   GraphicIOField "PlotLight_Round_G_33" at 416,264 size 24x24; PictureOn "PilotLight_Round_G_On_256c"; PictureOff "PilotLight_Round_G_Off_256c"
      ProcessValue <- "Senzor 2 proximitate softstarter aer destacker"

screen "Manual.Stacker" 800x480, template "TemplateWithClockAndBackBtnForManual"
   on GenerateScreen: SetBit("Maintenance")
   on ClearScreen: ResetBit("Maintenance")
   TextField "Text field_14" at 494,54 size 179x20; Text 'Comanda 1 softstarter aer'
   TextField "Text field_15" at 494,134 size 190x20; Text 'Comanda cilindru vertical jos'
   TextField "Text field_16" at 494,174 size 193x20; Text 'Comanda cilindru vertical sus'
   TextField "Text field_17" at 494,214 size 155x20; Text 'Comanda furca retrasa'
   TextField "Text field_18" at 494,254 size 153x20; Text 'Comanda furca extinsa'
   Switch "Switch_1" at 696,128 size 64x32; CaptionText 'Switch'; TextOff 'OFF'; TextOn 'ON'
      ProcessValue <- "S_Comanda cilindru vertical jos"
      on SwitchOn: SetBit("S_Comanda cilindru vertical jos")
      on SwitchOff: ResetBit("S_Comanda cilindru vertical jos")
   GraphicIOField "PlotLight_Round_G_2" at 160,48 size 24x24; PictureOff "PilotLight_Round_G_Off_256c"; PictureOn "PilotLight_Round_G_On_256c"
      ProcessValue <- "DB_PalletDispenser_PD2_Stacking_DB_PD1_MiddlePosition"
   TextField "Text field_3" at 16,50 size 126x20; Text 'PD1 MiddlePosition'
   Switch "Switch_2" at 696,48 size 64x32; CaptionText 'Switch'; TextOff 'OFF'; TextOn 'ON'
      ProcessValue <- "Comanda 1 softstarter aer stacker"
      on SwitchOn: SetBit("Comanda 1 softstarter aer stacker")
      on SwitchOff: ResetBit("Comanda 1 softstarter aer stacker")
   Switch "Switch_3" at 696,168 size 64x32; CaptionText 'Switch'; TextOff 'OFF'; TextOn 'ON'
      ProcessValue <- "S_Comanda cilindru vertical sus"
      on SwitchOn: SetBit("S_Comanda cilindru vertical sus")
      on SwitchOff: ResetBit("S_Comanda cilindru vertical sus")
   Switch "Switch_4" at 696,208 size 64x32; CaptionText 'Switch'; TextOff 'OFF'; TextOn 'ON'
      ProcessValue <- "S_Comanda furca retrasa"
      on SwitchOn: SetBit("S_Comanda furca retrasa")
      on SwitchOff: ResetBit("S_Comanda furca retrasa")
   Switch "Switch_5" at 696,248 size 64x32; CaptionText 'Switch'; TextOff 'OFF'; TextOn 'ON'
      ProcessValue <- "S_Comanda furca extinsa"
      on SwitchOn: SetBit("S_Comanda furca extinsa")
      on SwitchOff: ResetBit("S_Comanda furca extinsa")
   TextField "Text field_21" at 494,94 size 179x20; Text 'Comanda 2 softstarter aer'
   Switch "Switch_8" at 696,88 size 64x32; CaptionText 'Switch'; TextOff 'OFF'; TextOn 'ON'
      ProcessValue <- "Comanda 2 softstarter aer stacker"
      on SwitchOn: SetBit("Comanda 2 softstarter aer stacker")
      on SwitchOff: ResetBit("Comanda 2 softstarter aer stacker")
   GraphicIOField "PlotLight_Round_G_1" at 160,72 size 24x24; PictureOn "PilotLight_Round_G_On_256c"; PictureOff "PilotLight_Round_G_Off_256c"
      ProcessValue <- "DB_PalletDispenser_PD2_Stacking_DB_PD1_Up"
   TextField "Text field_1" at 16,74 size 50x20; Text 'PD1 Up'
   GraphicIOField "PlotLight_Round_G_3" at 160,96 size 24x24; PictureOn "PilotLight_Round_G_On_256c"; PictureOff "PilotLight_Round_G_Off_256c"
      ProcessValue <- "DB_PalletDispenser_PD2_Stacking_DB_PD1_Down"
   TextField "Text field_2" at 16,98 size 70x20; Text 'PD1 Down'
   GraphicIOField "PlotLight_Round_G_4" at 160,120 size 24x24; PictureOn "PilotLight_Round_G_On_256c"; PictureOff "PilotLight_Round_G_Off_256c"
      ProcessValue <- "DB_PalletDispenser_PD2_Stacking_DB_PD1_Forks_In"
   TextField "Text field_4" at 16,122 size 85x20; Text 'PD1 Forks In'
   GraphicIOField "PlotLight_Round_G_5" at 160,144 size 24x24; PictureOff "PilotLight_Round_G_Off_256c"; PictureOn "PilotLight_Round_G_On_256c"
      ProcessValue <- "DB_PalletDispenser_PD2_Stacking_DB_PD1_Forks_Out"
   TextField "Text field_5" at 16,146 size 95x20; Text 'PD1 Forks Out'
   GraphicIOField "PlotLight_Round_G_7" at 160,168 size 24x24; PictureOn "PilotLight_Round_G_On_256c"; PictureOff "PilotLight_Round_G_Off_256c"
      ProcessValue <- "DB_PalletDispenser_PD2_Stacking_DB_Alarm_Active"
   TextField "Text field_7" at 16,170 size 89x20; Text 'Alarm Active'
   GraphicIOField "PlotLight_Round_G_8" at 416,48 size 24x24; PictureOff "PilotLight_Round_G_Off_256c"; PictureOn "PilotLight_Round_G_On_256c"
      ProcessValue <- "S_Cilindru extins"
   TextField "Text field_8" at 240,50 size 111x20; Text 'S_Cilindru extins'
   GraphicIOField "PlotLight_Round_G_9" at 416,72 size 24x24; PictureOff "PilotLight_Round_G_Off_256c"; PictureOn "PilotLight_Round_G_On_256c"
      ProcessValue <- "S_Cilindru retras"
   TextField "Text field_9" at 240,74 size 113x20; Text 'S_Cilindru retras'
   GraphicIOField "PlotLight_Round_G_10" at 416,96 size 24x24; PictureOn "PilotLight_Round_G_On_256c"; PictureOff "PilotLight_Round_G_Off_256c"
      ProcessValue <- "S_Cilindru vertical jos"
   TextField "Text field_10" at 240,98 size 144x20; Text 'S_Cilindru vertical jos'
   GraphicIOField "PlotLight_Round_G_11" at 416,120 size 24x24; PictureOn "PilotLight_Round_G_On_256c"; PictureOff "PilotLight_Round_G_Off_256c"
      ProcessValue <- "S_Cilindru vertical mijloc"
   TextField "Text field_11" at 240,122 size 161x20; Text 'S_Cilindru vertical mijloc'
   GraphicIOField "PlotLight_Round_G_12" at 416,144 size 24x24; PictureOn "PilotLight_Round_G_On_256c"; PictureOff "PilotLight_Round_G_Off_256c"
      ProcessValue <- "S_Cilindru vertical sus"
   TextField "Text field_12" at 240,146 size 147x20; Text 'S_Cilindru vertical sus'
   GraphicIOField "PlotLight_Round_G_13" at 416,168 size 24x24; PictureOff "PilotLight_Round_G_Off_256c"; PictureOn "PilotLight_Round_G_On_256c"
      ProcessValue <- "S_Lungime 1"
   TextField "Text field_13" at 240,170 size 86x20; Text 'S_Lungime 1'
   GraphicIOField "PlotLight_Round_G_14" at 416,192 size 24x24; PictureOff "PilotLight_Round_G_Off_256c"; PictureOn "PilotLight_Round_G_On_256c"
      ProcessValue <- "S_Lungime 2"
   TextField "Text field_19" at 240,194 size 86x20; Text 'S_Lungime 2'
   GraphicIOField "PlotLight_Round_G_15" at 416,216 size 24x24; PictureOn "PilotLight_Round_G_On_256c"; PictureOff "PilotLight_Round_G_Off_256c"
      ProcessValue <- "S_Lungime 3"
   TextField "Text field_20" at 240,218 size 86x20; Text 'S_Lungime 3'
   GraphicIOField "PlotLight_Round_G_6" at 416,240 size 24x24; PictureOff "PilotLight_Round_G_Off_256c"; PictureOn "PilotLight_Round_G_On_256c"
      ProcessValue <- "S_Detectie palet"
   TextField "Text field_6" at 240,242 size 113x20; Text 'S_Detectie palet'
   GraphicIOField "PlotLight_Round_G_30" at 416,264 size 24x24; PictureOn "PilotLight_Round_G_On_256c"; PictureOff "PilotLight_Round_G_Off_256c"
      ProcessValue <- "Senzor 1 proximitate softstarter aer stacker"
   TextField "Text field_31" at 112,266 size 296x20; Text 'Senzor 1 proximitate softstarter aer stacker'
   GraphicIOField "PlotLight_Round_G_34" at 416,288 size 24x24; PictureOn "PilotLight_Round_G_On_256c"; PictureOff "PilotLight_Round_G_Off_256c"
      ProcessValue <- "Senzor 2 proximitate softstarter aer stacker"
   TextField "Text field_35" at 112,290 size 296x20; Text 'Senzor 2 proximitate softstarter aer stacker'

Template "TemplateWithClock" 800x480
   DateTimeField "Template_Date/time field_1" at 624,10 size 172x21
   GraphicView "Template_Graphic view_1" at 592,384 size 208x96; Picture "energom logo gonzales_1"

Template "TemplateWithClockAndBackBtn" 800x480
   Button "SB_NavigateLeft_48x48" at 72,0 size 64x40; TextOff 'Text'; PictureOff "SB_NavigateLeft_48x48_256c"
      on Press: function_efd93a16()
   Button "SB_NavigateHome_48x48" at 0,0 size 64x40; TextOff 'Text'; PictureOff "SB_NavigateHome_48x48_256c"
      on Press: ActivateScreen("Main", 0)
   DateTimeField "Template_Date/time field_1" at 624,10 size 172x21
   GraphicView "Template_Graphic view_1" at 592,384 size 208x96; Picture "energom logo gonzales_1"

Template "TemplateWithClockAndBackBtnForStatistics" 800x480
   Button "SB_NavigateHome_48x48" at 0,0 size 64x40; TextOff 'Text'; PictureOff "SB_NavigateHome_48x48_256c"
      on Press: ActivateScreen("Main", 0)
   Button "Button_4" at 8,392 size 136x80; TextOff 'Paleti Reparati'; Authorization "Operate"
      on Press: ActivateScreen("Production.Repair", 0); SetTag("CurrentScreenStatistics", 0)
      Visibility <- "CurrentUserGroup"
      Appearance <- "CurrentScreenStatistics"
   Button "Button_1" at 152,392 size 136x80; TextOff 'Paleti Demontati'; Authorization "Operate"
      on Press: ActivateScreen("Production.Destroy", 0); SetTag("CurrentScreenStatistics", 1)
      Visibility <- "CurrentUserGroup"
      Appearance <- "CurrentScreenStatistics"
   Button "Button_2" at 296,392 size 136x80; TextOff 'Energie'; Authorization "Operate"
      on Press: ActivateScreen("Energy", 0); SetTag("CurrentScreenStatistics", 2)
      Visibility <- "CurrentUserGroup"
      Appearance <- "CurrentScreenStatistics"
   Button "Button_3" at 440,392 size 136x80; TextOff 'Protectii'; Authorization "Operate"
      on Press: ActivateScreen("Safety", 0); SetTag("CurrentScreenStatistics", 3)
      Visibility <- "CurrentUserGroup"
      Appearance <- "CurrentScreenStatistics"
   DateTimeField "Template_Date/time field_1" at 624,10 size 172x21
   GraphicView "Template_Graphic view_1" at 592,384 size 208x96; Picture "energom logo gonzales_1"

Template "TemplateWithClockAndBackBtnForManual" 800x480
   Button "SB_NavigateHome_48x48" at 0,0 size 64x40; TextOff 'Text'; PictureOff "SB_NavigateHome_48x48_256c"
      on Press: ActivateScreen("Main", 0)
   DateTimeField "Template_Date/time field_1" at 624,10 size 172x21
   Button "Button_5" at 8,392 size 136x36; TextOff 'General'; Authorization "Operate"
      on Press: ActivateScreen("Manual.General", 0); SetTag("CurrentScreenManual", 0)
      Visibility <- "CurrentUserGroup"
      Appearance <- "CurrentScreenManual"
   Button "Button_6" at 152,392 size 136x36; TextOff 'Destacker'; Authorization "Operate"
      on Press: ActivateScreen("Manual.Destacker", 0); SetTag("CurrentScreenManual", 2)
      Visibility <- "CurrentUserGroup"
      Appearance <- "CurrentScreenManual"
   Button "Button_7" at 296,392 size 136x36; TextOff 'Stacker'; Authorization "Operate"
      on Press: ActivateScreen("Manual.Stacker", 0); SetTag("CurrentScreenManual", 4)
      Visibility <- "CurrentUserGroup"
      Appearance <- "CurrentScreenManual"
   Button "Button_8" at 8,436 size 136x36; TextOff 'Safety'; Authorization "Operate"
      on Press: ActivateScreen("Manual.Safety", 0); SetTag("CurrentScreenManual", 1)
      Visibility <- "CurrentUserGroup"
      Appearance <- "CurrentScreenManual"
   Button "Button_1" at 440,392 size 136x36; TextOff 'Transfer'; Authorization "Operate"
      on Press: ActivateScreen("Manual.Transfer", 0); SetTag("CurrentScreenManual", 6)
      Visibility <- "CurrentUserGroup"
      Appearance <- "CurrentScreenManual"
   GraphicView "Template_Graphic view_1" at 592,384 size 208x96; Picture "energom logo gonzales_1"
   Button "Button_2" at 152,436 size 136x36; TextOff 'Conveioare Destacker'; Authorization "Operate"
      on Press: ActivateScreen("Manual.DestackerConveyors", 0); SetTag("CurrentScreenManual", 3)
      Visibility <- "CurrentUserGroup"
      Appearance <- "CurrentScreenManual"
   Button "Button_3" at 296,436 size 136x36; TextOff 'Conveioare Stacker'; Authorization "Operate"
      on Press: ActivateScreen("Manual.StackerConveyors", 0); SetTag("CurrentScreenManual", 5)
      Visibility <- "CurrentUserGroup"
      Appearance <- "CurrentScreenManual"
   Button "Button_4" at 440,436 size 136x36; TextOff 'Diagnoza IO Link'; Authorization "Operate"
      on Press: ActivateScreen("Manual.IOLinkDiag", 0); SetTag("CurrentScreenManual", 7)
      Visibility <- "CurrentUserGroup"
      Appearance <- "CurrentScreenManual"

scheduled task "ChangeUserTask"
   on Action: function_f41c6f6c("CurrentUser"); function_e1ab61de("CurrentUserGroup"); function_de9337da()
*)

(* ===== HMI "HMI_RT_1" =====

graphic list "List": 1 'Graphic_4'; 2 'Graphic_6'; 4..16 'Graphic_7'

ScreenModuleEditorView "Transfer Paleta" 640x480
   GraphicIOField "Graphic I/O field_1" at 1,3 size 40x40; PictureList "List"
      ProcessValue <- "Step"
   GraphicView "Graphic view_1" at 11,13 size 20x20; Picture "Graphic_5"
      Visibility <- "Error"
*)

(* ===== HMI "HMI_RT_2" =====
system functions are stored by id; their names below are inferred from use
connection "HMI_Connection_2": ETHERNET, SMART_S7_1200_OMS

HMI tags "Default tag table"
   "Emergency Stop Stacker" : Bool = PLC 113S1 AT %I1.0, 1 s
   "Avarie Conveior 4 stacker" : Bool = PLC 128U1_Fault AT %I5.1, 1 s
   "Prezenta aer" : Bool = PLC 151S1 AT %I2.0, 1 s
   "Protectie cuplata Conveior 1 alimentare destacker" : Bool = PLC 120Q1 AT %I2.2, 1 s
   "Protectie cuplata Conveior 2 iesire destacker" : Bool = PLC 122Q1 AT %I2.7, 1 s
   "Avarie Conveior 1 alimentare destacker" : Bool = PLC 120U1_Fault AT %I2.6, 1 s
   "Avarie Conveior 2 iesire destacker" : Bool = PLC 122U1_Fault AT %I3.3, 1 s
   "Contactor cuplat Conveior 1 alimentare destacker" : Bool = PLC 121K1 AT %I2.3, 1 s
   "Contactor cuplat Conveior 2 iesire destacker" : Bool = PLC 123K1 AT %I3.0, 1 s
   "Frana decuplata Conveior 1 alimentare destacker" : Bool = PLC 120K1 AT %I2.4, 1 s
   "Frana decuplata Conveior 2 iesire destacker" : Bool = PLC 122K1 AT %I3.1, 1 s
   "Functionare Conveior 1 alimentare destacker" : Bool = PLC 120U1_PowerOK AT %I2.5, 1 s
   "Functionare Conveior 2 iesire destacker" : Bool = PLC 122U1_PowerOK AT %I3.2, 1 s
   "Senzor 1 proximitate softstarter aer destacker" : Bool = PLC 142VFA1_SQ1 AT %I6.4, 1 s
   "Senzor 2 proximitate softstarter aer destacker" : Bool = PLC 142VFA1_SQ2 AT %I6.5, 1 s
   "Reset safety Stacker_New" : Bool = PLC 1XXS2 AT %I68.6, 1 s
   "Comanda 1 softstarter aer destacker" : Bool = PLC "Comanda 1 softstarter aer stacker_new" AT %Q64.1, 1 s
   "Cuplare contactor VFD Conveior 1 alimentare destacker" : Bool = PLC CSN3_PowerOK AT %Q7.3, 1 s
   "Fault Aknowledge VFD Conveior 1 alimentare destacker" : Bool = PLC CSN3_FaultAck AT %Q10.0, 1 s
   "ON/OFF1 VFD Conveior 1 alimentare destacker" : Bool = PLC CSN3_Start AT %Q7.4, 1 s
   "Cuplare contactor VFD Conveior 2 iesire destacker" : Bool = PLC CSN4_PowerOK AT %Q7.5, 1 s
   "Fault Aknowledge VFD Conveior 2 iesire destacker" : Bool = PLC CSN4_FaultAck AT %Q10.1, 1 s
   "ON/OFF1 VFD Conveior 2 iesire destacker" : Bool = PLC CSN4_Start AT %Q7.6, 1 s
   "Contactor cuplat Conveior 4 descarcare stacker" : Bool = PLC 129K1 AT %I4.6, 1 s
   "Frana decuplata Conveior 4 descarcare stacker" : Bool = PLC 128K1 AT %I4.7, 1 s
   "Functionare Conveior 4 stacker" : Bool = PLC 128U1_PowerOK AT %I5.0, 1 s
   "Protectie cuplata Conveior 4 descarcare stacker" : Bool = PLC 128Q1 AT %I4.5, 1 s
   "Cuplare contactor VFD Conveior 4 descarcare stacker" : Bool = PLC CS4_PowerOK AT %Q8.5, 1 s
   "Fault Aknowledge VFD Conveior 4 descarcare stacker" : Bool = PLC CS4_FaultAck AT %Q10.3, 1 s
   "ON/OFF1 VFD Conveior 4 descarcare stacker" : Bool = PLC CS4_Start AT %Q8.6, 1 s
   "Avarie Conveior 3 transfer palet 2" : Bool = PLC 126U1_Fault AT %I4.4, 1 s
   "Contactor cuplat Conveior 3 transfer palet 2" : Bool = PLC 127K1 AT %I4.1, 1 s
   "Frana decuplata Conveior 3 transfer palet 2" : Bool = PLC 126K1 AT %I4.2, 1 s
   "Functionare Conveior 1 preluare paleti OK" : Bool = PLC 124K1 AT %I3.5, 1 s
   "Functionare Conveior 2 transfer palet 1" : Bool = PLC 125K1 AT %I3.7, 1 s
   "Functionare Conveior 3 transfer palet 2" : Bool = PLC 126U1_PowerOK AT %I4.3, 1 s
   "Protectie cuplata Conveior 1 preluare paleti OK" : Bool = PLC 124Q1 AT %I3.4, 1 s
   "Protectie cuplata Conveior 2 transfer palet 1" : Bool = PLC 125Q1 AT %I3.6, 1 s
   "Protectie cuplata Conveior 3 transfer palet 2" : Bool = PLC 126Q1 AT %I4.0, 1 s
   "Cuplare contactor VFD Conveior 3 transfer palet 2" : Bool = PLC CS3_PowerOK AT %Q8.3, 1 s
   "Fault Aknowledge VFD Conveior 3 transfer palet 2" : Bool = PLC CS3_FaultAck AT %Q10.2, 1 s
   "ON/OFF1 VFD Conveior 3 transfer palet 2" : Bool = PLC CS3_Start AT %Q8.4, 1 s
   "Softstarter aer 1.1 Conveior 1 preluare paleti OK" : Bool = PLC "Softstarter aer 1.1 Conveior 1 preluare paleti OK" AT %Q8.1, 1 s
   "Softstarter aer 1.2 Conveior 1 preluare paleti OK" : Bool = PLC "Softstarter aer 1.2 Conveior 1 preluare paleti OK" AT %Q8.2, 1 s
   "Start Conveior 1 preluare paleti OK" : Bool = PLC CS1_Start AT %Q8.0, 1 s
   "Start Conveior 2 transfer palet 1" : Bool = PLC CS2_Start AT %Q7.0, 1 s
   "Comanda 2 softstarter aer destacker" : Bool = PLC "Comanda 2 softstarter aer stacker_new" AT %Q66.1, 1 s
   "Comanda 1 softstarter aer stacker" : Bool = PLC "Comanda 1 softstarter aer stacker" AT %Q72.1, 1 s
   "Comanda 2 softstarter aer stacker" : Bool = PLC "Comanda 2 softstarter aer stacker" AT %Q74.1, 1 s
   "MD_IS1_SC_X1.0" : Bool = PLC "MD_IS1_SC_X1.0" AT %I70.0, 1 s
   "MD_IS1_SC_X1.1" : Bool = PLC "MD_IS1_SC_X1.1" AT %I70.1, 1 s
   "MD_IS1_SC_X1.2" : Bool = PLC "MD_IS1_SC_X1.2" AT %I70.2, 1 s
   "MD_IS1_SC_X1.3" : Bool = PLC "MD_IS1_SC_X1.3" AT %I70.3, 1 s
   "MD_IS1_SC_X1.4" : Bool = PLC "MD_IS1_SC_X1.4" AT %I70.4, 1 s
   "MD_IS1_SC_X1.5" : Bool = PLC "MD_IS1_SC_X1.5" AT %I70.5, 1 s
   "MD_IS1_SC_X1.6" : Bool = PLC "MD_IS1_SC_X1.6" AT %I70.6, 1 s
   "MD_IS1_SC_X1.7" : Bool = PLC "MD_IS1_SC_X1.7" AT %I70.7, 1 s
   "MD_IS2_SC_X1.0" : Bool = PLC "MD_IS2_SC_X1.0" AT %I75.0, 1 s
   "MD_IS2_SC_X1.1" : Bool = PLC "MD_IS2_SC_X1.1" AT %I75.1, 1 s
   "MD_IS2_SC_X1.2" : Bool = PLC "MD_IS2_SC_X1.2" AT %I75.2, 1 s
   "MD_IS2_SC_X1.3" : Bool = PLC "MD_IS2_SC_X1.3" AT %I75.3, 1 s
   "MD_IS2_SC_X1.4" : Bool = PLC "MD_IS2_SC_X1.4" AT %I75.4, 1 s
   "MD_IS2_SC_X1.5" : Bool = PLC "MD_IS2_SC_X1.5" AT %I75.5, 1 s
   "MD_IS2_SC_X1.6" : Bool = PLC "MD_IS2_SC_X1.6" AT %I75.6, 1 s
   "MD_IS2_SC_X1.7" : Bool = PLC "MD_IS2_SC_X1.7" AT %I75.7, 1 s
   "MD_OS_SC_X1.0" : Bool = PLC "MD_OS_SC_X1.0" AT %I92.0, 1 s
   "MD_OS_SC_X1.1" : Bool = PLC "MD_OS_SC_X1.1" AT %I93.0, 1 s
   "MD_OS_SC_X1.2" : Bool = PLC "MD_OS_SC_X1.2" AT %I92.1, 1 s
   "MD_OS_SC_X1.3" : Bool = PLC "MD_OS_SC_X1.3" AT %I93.1, 1 s
   "MD_OS_SC_X1.4" : Bool = PLC "MD_OS_SC_X1.4" AT %I92.2, 1 s
   "MD_OS_SC_X1.5" : Bool = PLC "MD_OS_SC_X1.5" AT %I93.2, 1 s
   "MS_IS1_SC_X1.0" : Bool = PLC "MS_IS1_SC_X1.0" AT %I80.0, 1 s
   "MS_IS1_SC_X1.1" : Bool = PLC "MS_IS1_SC_X1.1" AT %I80.1, 1 s
   "MS_IS1_SC_X1.2" : Bool = PLC "MS_IS1_SC_X1.2" AT %I80.2, 1 s
   "MS_IS1_SC_X1.3" : Bool = PLC "MS_IS1_SC_X1.3" AT %I80.3, 1 s
   "MS_IS1_SC_X1.4" : Bool = PLC "MS_IS1_SC_X1.4" AT %I80.4, 1 s
   "MS_IS1_SC_X1.5" : Bool = PLC "MS_IS1_SC_X1.5" AT %I80.5, 1 s
   "MS_IS1_SC_X1.6" : Bool = PLC "MS_IS1_SC_X1.6" AT %I80.6, 1 s
   "MS_IS1_SC_X1.7" : Bool = PLC "MS_IS1_SC_X1.7" AT %I80.7, 1 s
   "MS_IS2_SC_X1.0" : Bool = PLC "MS_IS2_SC_X1.0" AT %I85.0, 1 s
   "MS_IS2_SC_X1.1" : Bool = PLC "MS_IS2_SC_X1.1" AT %I85.1, 1 s
   "MS_IS2_SC_X1.2" : Bool = PLC "MS_IS2_SC_X1.2" AT %I85.2, 1 s
   "MS_IS2_SC_X1.3" : Bool = PLC "MS_IS2_SC_X1.3" AT %I85.3, 1 s
   "MS_IS2_SC_X1.4" : Bool = PLC "MS_IS2_SC_X1.4" AT %I85.4, 1 s
   "MS_IS2_SC_X1.5" : Bool = PLC "MS_IS2_SC_X1.5" AT %I85.5, 1 s
   "MS_IS2_SC_X1.6" : Bool = PLC "MS_IS2_SC_X1.6" AT %I85.6, 1 s
   "MS_IS2_SC_X1.7" : Bool = PLC "MS_IS2_SC_X1.7" AT %I85.7, 1 s
   "MS_OS_SC_X1.0" : Bool = PLC "MS_OS_SC_X1.0" AT %I101.0, 1 s
   "MS_OS_SC_X1.1" : Bool = PLC "MS_OS_SC_X1.1" AT %I102.0, 1 s
   "MS_OS_SC_X1.2" : Bool = PLC "MS_OS_SC_X1.2" AT %I101.1, 1 s
   "MS_OS_SC_X1.3" : Bool = PLC "MS_OS_SC_X1.3" AT %I102.1, 1 s
   "MS_OS_SC_X1.4" : Bool = PLC "MS_OS_SC_X1.4" AT %I101.2, 1 s
   "MS_OS_SC_X1.5" : Bool = PLC "MS_OS_SC_X1.5" AT %I102.2, 1 s
   "DS_Comanda cilindru vertical jos" : Bool = PLC "SN_Comanda cilindru vertical jos" AT %Q66.0, 1 s
   "DS_Comanda cilindru vertical sus" : Bool = PLC "SN_Comanda cilindru vertical sus" AT %Q64.0, 1 s
   "DS_Comanda furca retrasa" : Bool = PLC "SN_Comanda furca retrasa" AT %Q65.0, 1 s
   "DB_PalletDispenser_PD2_De_Stacking_DB_PD1_MiddlePosition" : Bool = PLC DB_PalletDispenser_PD2_Stacking_New_DB.PD1.MiddlePosition, 1 s
   "DB_PalletDispenser_PD2_De_Stacking_DB_PD1_Up" : Bool = PLC DB_PalletDispenser_PD2_Stacking_New_DB.PD1.Up, 1 s
   "DB_PalletDispenser_PD2_De_Stacking_DB_PD1_Down" : Bool = PLC DB_PalletDispenser_PD2_Stacking_New_DB.PD1.Down, 1 s
   "DB_PalletDispenser_PD2_De_Stacking_DB_PD1_Forks_In" : Bool = PLC DB_PalletDispenser_PD2_Stacking_New_DB.PD1.Forks_In, 1 s
   "DB_PalletDispenser_PD2_De_Stacking_DB_PD1_Forks_Out" : Bool = PLC DB_PalletDispenser_PD2_Stacking_New_DB.PD1.Forks_Out, 1 s
   "DB_PalletDispenser_PD2_De_Stacking_DB_Alarm_Active" : Bool = PLC DB_PalletDispenser_PD2_Stacking_New_DB.Alarm.Active, 1 s
   "DB_PalletDispenser_PD2_Stacking_DB_PD1_MiddlePosition" : Bool = PLC DB_PalletDispenser_PD2_Stacking_DB.PD1.MiddlePosition, 1 s
   "DB_PalletDispenser_PD2_Stacking_DB_PD1_Up" : Bool = PLC DB_PalletDispenser_PD2_Stacking_DB.PD1.Up, 1 s
   "DB_PalletDispenser_PD2_Stacking_DB_PD1_Down" : Bool = PLC DB_PalletDispenser_PD2_Stacking_DB.PD1.Down, 1 s
   "DB_PalletDispenser_PD2_Stacking_DB_PD1_Forks_In" : Bool = PLC DB_PalletDispenser_PD2_Stacking_DB.PD1.Forks_In, 1 s
   "DB_PalletDispenser_PD2_Stacking_DB_PD1_Forks_Out" : Bool = PLC DB_PalletDispenser_PD2_Stacking_DB.PD1.Forks_Out, 1 s
   "DB_PalletDispenser_PD2_Stacking_DB_Alarm_Active" : Bool = PLC DB_PalletDispenser_PD2_Stacking_DB.Alarm.Active, 1 s
   "S_Comanda cilindru vertical jos" : Bool = PLC "S_Comanda cilindru vertical jos" AT %Q74.0, 1 s
   "S_Comanda cilindru vertical sus" : Bool = PLC "S_Comanda cilindru vertical sus" AT %Q72.0, 1 s
   "S_Comanda furca retrasa" : Bool = PLC "S_Comanda furca retrasa" AT %Q73.0, 1 s
   "S_Comanda furca extinsa" : Bool = PLC "S_Comanda furca extinsa" AT %Q75.0, 1 s
   "Destacker 110KF1 Safety Relay" : Bool = PLC 110KF1 AT %I0.0, 1 s
   "Destacker 111KF1 Safety Barrier Relay" : Bool = PLC 111KF1 AT %I0.1, 1 s
   "Emergency Stop Destacker" : Bool = PLC 110S1 AT %I0.6, 1 s
   "Emergency Stop Zone 2" : Bool = PLC 112S1 AT %I0.7, 1 s
   "Stacker 113KF1 Safety Relay" : Bool = PLC 113KF1 AT %I0.3, 1 s
   "Stacker 114KF1 Safety Barrier Relay 1" : Bool = PLC 114KF1 AT %I0.4, 1 s
   "Stacker 115KF1 Safety Barrier Relay 2" : Bool = PLC 115KF1 AT %I0.5, 1 s
   "Zone 2 112KF1 Safety Relay" : Bool = PLC 112KF1 AT %I0.2, 1 s
   "Reset Stacker_New 110KF1 Safety Relay" : Bool = PLC 153K1 AT %Q0.0, 1 s
   "Reset Stacker_New 111KF1 Safety Barrier Relay" : Bool = PLC 153K2 AT %Q0.1, 1 s
   "Reset safety Zone 2" : Bool = PLC 155S1 AT %I1.1, 1 s
   "Reset Stacker 113KF1 Safety Relay" : Bool = PLC 153K4 AT %Q0.3, 1 s
   "Reset Stacker 114KF1 Safety Barrier Relay 1" : Bool = PLC 153K5 AT %Q0.4, 1 s
   "Reset Stacker 115KF1 Safety Barrier Relay 2" : Bool = PLC 153K6 AT %Q0.5, 1 s
   "Reset Zone 2 112KF1 Safety Relay" : Bool = PLC 153K3 AT %Q0.2, 1 s
   "FB_AlarmCounter_DB_Counters_Destacker 110KF1 Safety Relay_CV" : Int = PLC FB_AlarmCounter_DB.Counters."Destacker 110KF1 Safety Relay".CV, 1 s
   "FB_AlarmCounter_DB_Counters_Destacker 111KF1 Safety Barrier Relay_CV" : Int = PLC FB_AlarmCounter_DB.Counters."Destacker 111KF1 Safety Barrier Relay".CV, 1 s
   "FB_AlarmCounter_DB_Counters_Zone 2 112KF1 Safety Relay_CV" : Int = PLC FB_AlarmCounter_DB.Counters."Zone 2 112KF1 Safety Relay".CV, 1 s
   "FB_AlarmCounter_DB_Counters_Stacker 113KF1 Safety Relay_CV" : Int = PLC FB_AlarmCounter_DB.Counters."Stacker 113KF1 Safety Relay".CV, 1 s
   "FB_AlarmCounter_DB_Counters_Stacker 114KF1 Safety Barrier Relay 1_CV" : Int = PLC FB_AlarmCounter_DB.Counters."Stacker 114KF1 Safety Barrier Relay 1".CV, 1 s
   "FB_AlarmCounter_DB_Counters_Stacker 115KF1 Safety Barrier Relay 2_CV" : Int = PLC FB_AlarmCounter_DB.Counters."Stacker 115KF1 Safety Barrier Relay 2".CV, 1 s
   "FB_AlarmCounter_DB_Counters_Emergency Stop Destacker_CV" : Int = PLC FB_AlarmCounter_DB.Counters."Emergency Stop Destacker".CV, 1 s
   "FB_AlarmCounter_DB_Counters_Emergency Stop Zone 2_CV" : Int = PLC FB_AlarmCounter_DB.Counters."Emergency Stop Zone 2".CV, 1 s
   "FB_AlarmCounter_DB_Counters_Emergency Stop Stacker_CV" : Int = PLC FB_AlarmCounter_DB.Counters."Emergency Stop Stacker".CV, 1 s
   "FB_EnergyCounter_DB_Counters_LastHour_CV" : UInt = PLC FB_EnergyCounter_DB.Counters.LastHour.CV, 1 s
   "FB_EnergyCounter_DB_Counters_LastDay_CV" : UDInt = PLC FB_EnergyCounter_DB.Counters.LastDay.CV, 1 s
   "FB_EnergyCounter_DB_Counters_LastMonth_CV" : UDInt = PLC FB_EnergyCounter_DB.Counters.LastMonth.CV, 1 s
   "Aliniere palet" : Bool = PLC CSN1_SQ3 AT %I68.1, 1 s
   "Centror extins" : Bool = PLC CP2_SQ3 AT %I79.5, 1 s
   "Centror retras" : Bool = PLC CP2_SQ2 AT %I78.5, 1 s
   "Detectie palet" : Bool = PLC "SN_Detectie palet" AT %I73.4, 1 s
   "DS_Cilindru extins" : Bool = PLC "SN_Cilindru extins" AT %I74.6, 1 s
   "DS_Cilindru retras" : Bool = PLC "SN_Cilindru retras" AT %I74.1, 1 s
   "DS_Cilindru vertical jos" : Bool = PLC "SN_Cilindru vertical jos" AT %I73.5, 1 s
   "DS_Cilindru vertical mijloc" : Bool = PLC "SN_Cilindru vertical mijloc" AT %I73.3, 1 s
   "DS_Cilindru vertical sus" : Bool = PLC "SN_Cilindru vertical sus" AT %I73.2, 1 s
   "DS_Lungime 1" : Bool = PLC CSN3_SQ2 AT %I68.3, 1 s
   "DS_Lungime 2" : Bool = PLC CSN3_SQ3 AT %I69.3, 1 s
   "DS_Lungime 3" : Bool = PLC CSN4_SQ1 AT %I68.4, 1 s
   "Feed palet" : Bool = PLC SN_Prez_conveyor_volum AT %I69.6, 1 s
   "Masurare lungime" : Bool = PLC CS2_SQ1 AT %I78.2, 1 s
   "Prezenta palet iesire" : Bool = PLC SN_Switch_Iesire AT %I69.4, 1 s
   "Prezenta palet_capat_conveyor" : Bool = PLC CS1_SQ3 AT %I78.1, 1 s
   "Prezenta palet_centror" : Bool = PLC "S_Prezenta palet_centror" AT %I79.1, 1 s
   "Prezenta palet_stanga" : Bool = PLC CS1_SQ1 AT %I78.0, 1 s
   "Prezenta_stiva" : Bool = PLC CS4_SQ1 AT %I78.4, 1 s
   "Prezenta stiva" : Bool = PLC CSN1_SQ1 AT %I68.0, 1 s
   "Protectie cuplata Circular masa fixa" : Bool = PLC 104F1 AT %I5.4, 1 s
   "Protectie cuplata HMI" : Bool = PLC 149F1 AT %I7.0, 1 s
   "Protectie cuplata Iluminat" : Bool = PLC 105F2 AT %I2.1, 1 s
   "Protectie cuplata Masina demontare paleti dreapta" : Bool = PLC 103F1 AT %I5.3, 1 s
   "Protectie cuplata Masina demontare paleti stanga" : Bool = PLC 102F1 AT %I5.2, 1 s
   "Protectie cuplata Post reparatie stanga+dreapta" : Bool = PLC 105F1 AT %I5.5, 1 s
   "Protectie cuplata Post reparatii minore" : Bool = PLC 106F1 AT %I5.6, 1 s
   "Protectie cuplata TELE" : Bool = PLC 107F1 AT %I5.7, 1 s
   "S_Cilindru extins" : Bool = PLC "S_Cilindru extins" AT %I84.6, 1 s
   "S_Cilindru retras" : Bool = PLC "S_Cilindru retras" AT %I84.1, 1 s
   "S_Cilindru vertical jos" : Bool = PLC "S_Cilindru vertical jos" AT %I83.5, 1 s
   "S_Cilindru vertical mijloc" : Bool = PLC "S_Cilindru vertical mijloc" AT %I83.3, 1 s
   "S_Cilindru vertical sus" : Bool = PLC "S_Cilindru vertical sus" AT %I83.2, 1 s
   "S_Lungime 1" : Bool = PLC CS3_SQ1 AT %I79.2, 1 s
   "S_Lungime 2" : Bool = PLC CS3_SQ2 AT %I78.3, 1 s
   "S_Lungime 3" : Bool = PLC CS3_SQ3 AT %I79.3, 1 s
   "S_Detectie palet" : Bool = PLC "S_Detectie palet" AT %I83.4, 1 s
   "Senzor 1 proximitate softstarter aer stacker" : Bool = PLC 143VFA1_SQ1 AT %I83.7, 1 s
   "Senzor 1 proximitate softstarter aer zona 2" : Bool = PLC 141VFA1_SQ1 AT %I7.1, 1 s
   "Senzor 2 proximitate softstarter aer stacker" : Bool = PLC 143VFA1_SQ2 AT %I84.7, 1 s
   "Senzor 2 proximitate softstarter aer zona 2" : Bool = PLC 141VFA1_SQ2 AT %I7.2, 1 s
   "Senzor destacking" : Bool = PLC "SN_Senzor stacking" AT %I73.1, 1 s
   "Senzor stacking" : Bool = PLC "S_Senzor stacking" AT %I83.1, 1 s
   "Start masurare lungime" : Bool = PLC CSN3_SQ1 AT %I69.2, 1 s
   "DS_Comanda furca extinsa" : Bool = PLC "SN_Comanda furca extinsa" AT %Q67.0, 1 s
   "DB20_DATA_HMI_Step_Destacker" : Int = PLC DB20_DATA_HMI.Step_Destacker, 1 s
   "DB20_DATA_HMI_Step_Stacker" : Int = PLC DB20_DATA_HMI.Step_Stacker, 1 s
   "Maintenance" : Bool = PLC Maintenance AT %M5.0, 1 s
   "Rez_G7_DS" : Bool = PLC Rez_G7_DS AT %M6.0, 1 s
   "Rez_G7_S" : Bool = PLC Rez_G7_S AT %M6.1, 1 s
   "Fault_Length_DS" : Bool = PLC Fault_Length_DS AT %M6.2, 1 s
   "Fault_Length_DS_ACK" : Bool = PLC Fault_Length_DS_ACK AT %M6.4, 1 s
   "Length_DS_HMI_1" : Bool = PLC Length_DS_HMI_1 AT %M14.0, 1 s
   "Length_DS_HMI_2" : Bool = PLC Length_DS_HMI_2 AT %M14.1, 1 s
   "Length_DS_HMI_3" : Bool = PLC Length_DS_HMI_3 AT %M14.2, 1 s
   "Length_S_HMI_1" : Bool = PLC Length_S_HMI_1 AT %M14.3, 1 s
   "Length_S_HMI_2" : Bool = PLC Length_S_HMI_2 AT %M14.4, 1 s
   "Length_S_HMI_3" : Bool = PLC Length_S_HMI_3 AT %M14.5, 1 s
   "Fault_Length_S_ACK" : Bool = PLC Fault_Length_S_ACK AT %M6.5, 1 s
   "Fault_Length_S" : Bool = PLC Fault_Length_S AT %M6.3, 1 s
   "DB3_FAULTS_Alarm_Safety_SN" : Word = PLC DB3_FAULTS.Alarm_Safety_SN AT %DB3.DBW22, 1 s
   "DB3_FAULTS_Alarm_Safety_Z2" : Word = PLC DB3_FAULTS.Alarm_Safety_Z2 AT %DB3.DBW24, 1 s
   "DB3_FAULTS_Alarm_Safety_S" : Word = PLC DB3_FAULTS.Alarm_Safety_S AT %DB3.DBW26, 1 s
   "DB3_FAULTS_Alarm_CD1" : Word = PLC DB3_FAULTS.Alarm_CD1 AT %DB3.DBW10, 1 s
   "DB3_FAULTS_Alarm_CD2" : Word = PLC DB3_FAULTS.Alarm_CD2 AT %DB3.DBW12, 1 s
   "FB_ProductionStatistics_DB_Counters_Destroyed_LastDay_CV" : Int = PLC FB_ProductionStatistics_DB.Counters.Destroyed.LastDay.CV, 1 s
   "FB_ProductionStatistics_DB_Counters_Repairs_LastDay_CV" : Int = PLC FB_ProductionStatistics_DB.Counters.Repairs.LastDay.CV, 1 s
   "Manual_Comanda 1 softstarter aer destacker" : Bool = PLC "Manual_Comanda 1 softstarter aer destacker" AT %M11.1, 1 s
   "Manual_Comanda 2 softstarter aer destacker" : Bool = PLC "Manual_Comanda 2 softstarter aer destacker" AT %M11.2, 1 s
   "Manual_Cuplare contactor VFD Conveior 1 alimentare destacker" : Bool = PLC "Manual_Cuplare contactor VFD Conveior 1 alimentare destacker" AT %M8.6, 1 s
   "Manual_Fault Aknowledge VFD Conveior 1 alimentare destacker" : Bool = PLC "Manual_Fault Aknowledge VFD Conveior 1 alimentare destacker" AT %M9.0, 1 s
   "Manual_ON/OFF1 VFD Conveior 1 alimentare destacker" : Bool = PLC "Manual_ON/OFF1 VFD Conveior 1 alimentare destacker" AT %M8.7, 1 s
   "Manual_Cuplare contactor VFD Conveior 2 iesire destacker" : Bool = PLC "Manual_Cuplare contactor VFD Conveior 2 iesire destacker" AT %M9.1, 1 s
   "Manual_ON/OFF1 VFD Conveior 2 iesire destacker" : Bool = PLC "Manual_ON/OFF1 VFD Conveior 2 iesire destacker" AT %M9.2, 1 s
   "Manual_Reset Stacker_New 110KF1 Safety Relay" : Bool = PLC "Manual_Reset Destacker 110KF1 Safety Relay" AT %M8.0, 1 s
   "Manual_Reset Destacker 111KF1 Safety Barrier Relay" : Bool = PLC "Manual_Reset Destacker 111KF1 Safety Barrier Relay" AT %M8.1, 1 s
   "Manual_Reset Zone 2 112KF1 Safety Relay" : Bool = PLC "Manual_Reset Zone 2 112KF1 Safety Relay" AT %M8.2, 1 s
   "Manual_Reset Stacker 113KF1 Safety Relay" : Bool = PLC "Manual_Reset Stacker 113KF1 Safety Relay" AT %M8.3, 1 s
   "Manual_Reset Stacker 114KF1 Safety Barrier Relay 1" : Bool = PLC "Manual_Reset Stacker 114KF1 Safety Barrier Relay 1" AT %M8.4, 1 s
   "Manual_Reset Stacker 115KF1 Safety Barrier Relay 2" : Bool = PLC "Manual_Reset Stacker 115KF1 Safety Barrier Relay 2" AT %M8.5, 1 s
   "Manual_Comanda 1 softstarter aer stacker" : Bool = PLC "Manual_Comanda 1 softstarter aer stacker" AT %M12.0, 1 s
   "Manual_Comanda 2 softstarter aer stacker" : Bool = PLC "Manual_Comanda 2 softstarter aer stacker" AT %M12.1, 1 s
   "Manual_Cuplare contactor VFD Conveior 4 descarcare stacker" : Bool = PLC "Manual_Cuplare contactor VFD Conveior 4 descarcare stacker" AT %M10.3, 1 s
   "Manual_Fault Aknowledge VFD Conveior 4 descarcare stacker" : Bool = PLC "Manual_Fault Aknowledge VFD Conveior 4 descarcare stacker" AT %M10.5, 1 s
   "Manual_ON/OFF1 VFD Conveior 4 descarcare stacker" : Bool = PLC "Manual_ON/OFF1 VFD Conveior 4 descarcare stacker" AT %M10.4, 1 s
   "Manual_Cuplare contactor VFD Conveior 3 transfer palet 2" : Bool = PLC "Manual_Cuplare contactor VFD Conveior 3 transfer palet 2" AT %M10.0, 1 s
   "Manual_Fault Aknowledge VFD Conveior 3 transfer palet 2" : Bool = PLC "Manual_Fault Aknowledge VFD Conveior 3 transfer palet 2" AT %M10.2, 1 s
   "Manual_ON/OFF1 VFD Conveior 3 transfer palet 2" : Bool = PLC "Manual_ON/OFF1 VFD Conveior 3 transfer palet 2" AT %M10.1, 1 s
   "Manual_Softstarter aer 1.1 Conveior 1 preluare paleti OK" : Bool = PLC "Manual_Softstarter aer 1.1 Conveior 1 preluare paleti OK" AT %M9.5, 1 s
   "Manual_Softstarter aer 1.2 Conveior 1 preluare paleti OK" : Bool = PLC "Manual_Softstarter aer 1.2 Conveior 1 preluare paleti OK" AT %M9.6, 1 s
   "Manual_Start Conveior 1 preluare paleti OK" : Bool = PLC "Manual_Start Conveior 1 preluare paleti OK" AT %M9.4, 1 s
   "Manual_Start Conveior 2 transfer palet 1" : Bool = PLC "Manual_Start Conveior 2 transfer palet 1" AT %M9.7, 1 s
   "Manual_DS" : Bool = PLC Manual_DS AT %M13.2, 1 s
   "Manual_S" : Bool = PLC Manual_S AT %M15.1, 1 s
   "s_f{1}_HMI_stat_s" : USInt = PLC s.f[1].HMI_statS, 1 s
   "s_f{1}_HMI_stat_t" : USInt = PLC s.f[1].HMI_statT, 1 s
   "ds_f{1}_HMI_stat_t" : USInt = PLC ds.f[1].HMI_statT, 1 s
   "s_f{4}_HMI_stat_s" : USInt = PLC s.f[4].HMI_statS, 1 s
   "s_f{2}_HMI_stat_s" : USInt = PLC s.f[2].HMI_statS, 1 s
   "s_f{3}_HMI_stat_s" : USInt = PLC s.f[3].HMI_statS, 1 s
   "s_f{3}_HMI_stat_t" : USInt = PLC s.f[3].HMI_statT, 1 s
   "ds_f{3}_HMI_stat_s" : USInt = PLC ds.f[1].HMI_statS, 1 s
   "s_f{2}_HMI_stat_t" : USInt = PLC s.f[2].HMI_statT, 1 s
   "s_f{5}_HMI_stat_s" : USInt = PLC s.f[5].HMI_statS, 1 s
   "s_f{4}_HMI_stat_t" : USInt = PLC s.f[4].HMI_statT, 1 s
   "ds_f{2}_HMI_stat_s" : USInt = PLC ds.f[1].HMI_statS, 1 s
   "ds_f{2}_HMI_stat_t" : USInt = PLC ds.f[1].HMI_statT, 1 s
   "ds_f{1}_HMI_stat_s" : USInt = PLC ds.f[1].HMI_statS, 1 s
   "O_Alm_Stack_Up" : Word = PLC O.S_Alm_Stack_Up AT %DB1.DBW0, 1 s
   "O_FurcaStacker_New_AlarmW" : Word = PLC O.FurcaStacker_New.AlarmW AT %DB1.DBW0, 1 s
   "O_CilindruVerticalStacker_New_AlarmW" : Word = PLC O.CilindruVerticalStacker_New.AlarmW AT %DB3.DBW2, 1 s
   "O_FurcaStacker_AlarmW" : Word = PLC O.FurcaStacker.AlarmW AT %DB1.DBX0.0, 1 s
   "Manual_S_Comanda cilindru vertical sus" : Bool = PLC O.CilindruVerticalStacker.ButAv AT %M11.4, 1 s
   "Manual_S_Comanda cilindru vertical jos" : Bool = PLC O.CilindruVerticalStacker.ButRet AT %M11.5, 1 s
   "Manual_S_Comanda furca extinsa" : Bool = PLC O.FurcaStacker.ButAv AT %M11.6, 1 s
   "Manual_DS_Comanda cilindru vertical jos" : Bool = PLC O.CilindruVerticalStacker_New.ButRet AT %M10.7, 1 s
   "Manual_DS_Comanda cilindru vertical sus" : Bool = PLC O.CilindruVerticalStacker_New.ButAv AT %M10.6, 1 s
   "Manual_DS_Comanda furca retrasa" : Bool = PLC O.FurcaStacker_New.ButRet AT %M11.0, 1 s
   "Manual_DS_Comanda furca extinsa" : Bool = PLC O.FurcaStacker_New.ButAv AT %M12.4, 1 s
   "Manual_S_Comanda centror extins" : Bool = PLC O.Centror_A.ButAv AT %DB1.DBX0.0, 1 s
   "O_CilindruVerticalStacker_StatRet" : USInt = PLC O.CilindruVerticalStacker.StatRet AT %DB1.DBX0.0, 1 s
   "O_CilindruVerticalStacker_New_StatRet" : USInt = PLC O.CilindruVerticalStacker_New.StatRet AT %DB1.DBB0, 1 s
   "O_FurcaStacker_StatAv" : USInt = PLC O.FurcaStacker.StatAv AT %DB1.DBB0, 1 s
   "O_FurcaStacker_New_StatAv" : USInt = PLC O.FurcaStacker_New.StatAv AT %DB1.DBB0, 1 s
   "O_FurcaStacker_StatRet" : USInt = PLC O.FurcaStacker.StatRet AT %DB1.DBB0, 1 s
   "O_Centror_StatAv" : USInt = PLC O.Centror_A.StatAv AT %DB1.DBB0, 1 s
   "O_CilindruVerticalStacker_New_StatAv" : USInt = PLC O.CilindruVerticalStacker_New.StatAv AT %DB1.DBB0, 1 s
   "O_Centror_StatRet" : USInt = PLC O.Centror_A.StatRet AT %DB1.DBB0, 1 s
   "Manual_S_Comanda centror retras" : Bool = PLC O.Centror_A.ButRet AT %DB1.DBX0.0, 1 s
   "O_CilindruVerticalStacker_StatAv" : USInt = PLC O.CilindruVerticalStacker.StatAv AT %DB1.DBX0.0, 1 s
   "O_FurcaStacker_New_StatRet" : USInt = PLC O.FurcaStacker_New.StatRet AT %DB1.DBB0, 1 s
   "bStop_S" : Bool = PLC bStop_S AT %M16.3, 1 s
   "bStart_S" : Bool = PLC bStart_S AT %M7.7, 1 s
   "bStop_DS" : Bool = PLC bStop_DS AT %M16.1, 1 s
   "bStepper_S" : Bool = PLC bStepper_S AT %M12.6, 1 s
   "bStepper_DS" : Bool = PLC bStepper_DS AT %M12.7, 1 s
   "bStart_DS" : Bool = PLC bStart_SN AT %M20.2, 1 s
   "forcep" : Bool = PLC ForceIniProdus AT %M7.6, 1 s
   "rsta" : Bool = PLC RstAlm AT %M7.4, 1 s
   "forcet" : Bool = PLC ForceIniTranzit AT %M7.5, 1 s
   "forcec" : Bool = PLC ForceIniCylRet AT %M17.0, 1 s
   "s_f{4}_AlarmW" : Word = PLC s.f[4].AlarmW AT %DB3.DBW18, 1 s
   "s_f{2}_AlarmW" : Word = PLC s.f[2].AlarmW AT %DB3.DBW14, 1 s
   "s_f{3}_AlarmW" : Word = PLC s.f[3].AlarmW AT %DB3.DBW16, 1 s
   "s_f{5}_AlarmW" : Word = PLC s.f[5].AlarmW AT %DB3.DBW20, 1 s
   "O_Centror_AlarmW" : Word = PLC O.Centror_A.AlarmW AT %DB3.DBW8, 1 s
   "s_f{1}_AlarmW" : Word = PLC s.f[1].AlarmW AT %DB1.DBB0, 1 s
   "Manual_S_Comanda furca retrasa" : Bool = PLC O.FurcaStacker.ButRet AT %M11.7, 1 s
   "DB3_FAULTS_Alarm_General" : Word = PLC DB3_FAULTS.Alarm_General_S AT %DB3.DBW28, 1 s
   "DB_MDM_S_Safe" : Bool = PLC DB_MDM_S.Safe, 1 s
   "DB_MDM_SN_step" : USInt = PLC DB_MDM_SN.step, 1 s
   "DB_MDM_S_step" : USInt = PLC DB_MDM_S.step, 1 s
   "Automat_DS" : Bool = PLC Automat_SN AT %M19.6, 1 s
   "Automat_S" : Bool = PLC Automat_S AT %M15.2, 1 s
   "O_Alm_Stack_Mid" : Word = PLC O.S_Alm_Stack_Mid AT %DB1.DBW0, 1 s
   "O_Alm_Stack_Dwn" : Word = PLC O.S_Alm_Stack_Dwn AT %DB1.DBW0, 1 s
   "inst_sel" : Int = PLC HMI.instance_sel AT %DB46.DBW42, 1 s
   "HMI.msop_viz" : USInt = PLC HMI.msop_vizi AT %DB46.DBB62, 1 s
   "numCyl" : USInt = PLC HMI.numCyl AT %DB46.DBB46, 1 s
   "numSens" : USInt = PLC HMI.numSens AT %DB46.DBB47, 1 s
   "numSt" : USInt = PLC HMI.numSt AT %DB46.DBB44, 1 s
   "numSt_s" : USInt = PLC HMI.numSt_s AT %DB46.DBB45, 1 s
   "pgCfg" : USInt = PLC HMI.pgCfg AT %DB46.DBB48, 1 s
   "ButOpW" : USInt = PLC HMI.ButOpHMI AT %DB46.DBB61, 1 s
   "ButOpMem" : USInt = PLC HMI.ButOpMem AT %DB46.DBB59, 1 s
   "ButOpVis" : USInt = PLC HMI.ButOpVis AT %DB46.DBB50, 1 s
   "butop_1" : Bool = PLC HMI.ButOp[1] AT %DB46.DBX52.1, 1 s
   "butop_2" : Bool = PLC HMI.ButOp[2] AT %DB46.DBX52.2, 1 s
   "butop_3" : Bool = PLC HMI.ButOp[3] AT %DB46.DBX52.3, 1 s
   "chg_prio" : Bool = PLC HMI.chg_prio AT %DB46.DBX58.0, 1 s
   "100KF1" : Bool = PLC 100KF1 AT %I1.3, 1 s
   "DB20_DATA_HMI_Reset_Faults" : Bool = PLC DB20_DATA_HMI.Reset_Faults, 1 s
   "DB3_FAULTS_Alarm_General_SN" : Word = PLC DB3_FAULTS.Alarm_General_SN AT %DB3.DBW30, 1 s
   "bStop_SN" : Bool = PLC bStop_SN AT %M20.1, 1 s
   "bStepper_SN" : Bool = PLC bStepper_SN AT %M20.0, 1 s
   "DB2_WORK_BITS_MDM{0}" : MDM = PLC DB2_WORK_BITS.MDM[0] AT %DB1.DBX0.0, 1 s
   "DB2_WORK_BITS_Select_MDM" : Int = PLC DB2_WORK_BITS.Select_MDM, 1 s
   "HMI_SN_msop_vizi" : USInt = PLC HMI_SN.msop_vizi AT %DB64.DBB62, 1 s
   "HMI_SN_numSt" : USInt = PLC HMI_SN.numSt AT %DB64.DBB44, 1 s
   "HMI_SN_numSt_s" : USInt = PLC HMI_SN.numSt_s AT %DB64.DBB45, 1 s
   "O_Centror_B_StatRet" : USInt = PLC O.Centror_B.StatRet, 1 s
   "O_Centror_B_StatAv" : USInt = PLC O.Centror_B.StatAv, 1 s
   "O_Centror_B_ButAv" : Bool = PLC O.Centror_B.ButAv, 1 s
   "O_Centror_B_ButRet" : Bool = PLC O.Centror_B.ButRet, 1 s

HMI tags "Alarms"
   "DS_AlarmMovement" : Word = PLC DS_AlarmMovement AT %MW2, 1 s
   "S_AlarmMovement" : Word = PLC S_AlarmMovement AT %MW4, 1 s

HMI tags "UserManagement"
   "CurrentUser" : WString[254], internal
   "CurrentUserGroup" : Int, internal

HMI tags "Statistics"
   "PalletsLastMonth" : Int, internal
   "PalletsLastWeek" : Int, internal
   "PalletsPerShift" : Array [0..8] of Int, internal

HMI tags "UI"
   "CurrentScreenStatistics" : Int, internal
   "CurrentScreenManual" : Bool = PLC DB20_DATA_HMI.Maintenance, 1 s
   "SwitchTestBit" : Bool, internal

HMI tags "status"
   "stS1" : Int, internal

discrete alarms
   40: 'Stiva nu a ajuns la stacker nou la timp', class Errors, trigger "DB3_FAULTS_Alarm_CD2" bit 0
   41: 'Paletul nu a ajuns la iesire la timp', class Errors, trigger "DB3_FAULTS_Alarm_CD2" bit 1
   42: 'Stiva nu a plecat spre stacker nou', class Errors, trigger "DB3_FAULTS_Alarm_CD1" bit 0
   43: 'Paletul nu a plecat de la stacker nou', class Errors, trigger "DB3_FAULTS_Alarm_CD2" bit 2
   44: 'Safety Linia B : Buton oprire urgenta apasat : <110KF1>', class Errors, trigger "DB3_FAULTS_Alarm_Safety_SN" bit 0
   46: 'Safety Linia A : Buton oprire urgenta apasat : <112KF1>', class Errors, trigger "DB3_FAULTS_Alarm_Safety_S" bit 0
   49: 'Safety Zona2A: Usa deschisa : <114KF1>', class Errors, trigger "DB3_FAULTS_Alarm_Safety_S" bit 2
   50: 'Safety Linia A : Bariera mutting stacker dezarmata <115KF1>', class Errors, trigger "DB3_FAULTS_Alarm_Safety_S" bit 3
   51: 'Safety Zona2B: Usa deschisa : <113KF1>', class Errors, trigger "DB3_FAULTS_Alarm_Safety_SN" bit 2
   52: 'Safety General : Usa principala deschisa : <100KF1>', class Errors, trigger "DB3_FAULTS_Alarm_Safety_S" bit 4
   21: 'Furca stacker nou a pierdut detectia in pozitia avans (4D; S1_B5)', class Errors, trigger "O_FurcaStacker_New_AlarmW" bit 2
   2: 'Alarma stacker nou miscare furci', class Errors, trigger "O_FurcaStacker_New_AlarmW" bit 7
   19: 'Furca stacker nou nu s-a retras in timpul prestabilit (4D; S1_B13)', class Errors, trigger "O_FurcaStacker_New_AlarmW" bit 4
   4: 'Alarma stacker miscare verticala', class Errors, trigger "O_FurcaStacker_AlarmW" bit 7
   10: 'Furca stacker nu a avansat in timpul prestabilit (4D; S1_B5)', class Errors, trigger "O_FurcaStacker_AlarmW" bit 0
   32: 'Palet aparut la postul de lucru fara transfer', class Errors, trigger "s_f{2}_AlarmW" bit 1
   33: 'Palet disparut de la postul de lucru fara transfer', class Errors, trigger "s_f{2}_AlarmW" bit 2
   29: 'Paletul nu a plecat de la postul de lucru', class Errors, trigger "s_f{2}_AlarmW" bit 0
   56: 'Palet disparut de la postul de lucru fara transfer', class Errors, trigger "s_f{1}_AlarmW" bit 2
   54: 'Paletul nu a plecat de la postul de lucru', class Errors, trigger "s_f{1}_AlarmW" bit 0
   55: 'Palet aparut la postul de lucru fara transfer', class Errors, trigger "s_f{1}_AlarmW" bit 1
   28: 'Stiva nu s-a evacuat la timp', class Errors, trigger "s_f{5}_AlarmW" bit 3
   26: 'Paletul nu a ajuns la centror la timp', class Errors, trigger "s_f{3}_AlarmW" bit 4
   36: 'Palet aparut la stacker fara transfer', class Errors, trigger "s_f{4}_AlarmW" bit 5
   30: 'Paletul nu a plecat de la centror', class Errors, trigger "s_f{3}_AlarmW" bit 5
   31: 'Stiva nu a plecat de la Stacker', class Errors, trigger "s_f{4}_AlarmW" bit 4
   38: 'Palet/Stiva aparut la evacuare fara transfer', class Errors, trigger "s_f{5}_AlarmW" bit 2
   27: 'Paletul nu a ajuns la stacker la timp', class Errors, trigger "s_f{4}_AlarmW" bit 3
   35: 'Palet disparut de la centror fara transfer', class Errors, trigger "s_f{3}_AlarmW" bit 3
   34: 'Palet aparut la centror fara transfer', class Errors, trigger "s_f{3}_AlarmW" bit 6
   37: 'Palet disparut de la stacker fara transfer', class Errors, trigger "s_f{4}_AlarmW" bit 2
   39: 'Palet/Stiva disparut de la evacuare fara transfer', class Errors, trigger "s_f{5}_AlarmW" bit 0
   8: 'Centrorul se afla in pozitia retras cu actionare (9D; CP2_SQ2)', class Errors, trigger "O_Centror_AlarmW" bit 1
   9: 'Centrorul a pierdut pozitia de avans (9D; CP2_SQ2)', class Errors, trigger "O_Centror_AlarmW" bit 2
   18: 'Furca stacker nou nu a avansat in timpul prestabilit (4D; S1_B5)', class Errors, trigger "O_FurcaStacker_New_AlarmW" bit 0
   12: 'Furca stacker blocata in pozitia de retras', class Errors, trigger "O_FurcaStacker_AlarmW" bit 1
   13: 'Furca stacker a pierdut detectia in pozitia avans (4D; S1_B5)', class Errors, trigger "O_FurcaStacker_AlarmW" bit 2
   7: 'Centrorul nu a realizat miscarea avans in timpul prestabilit (9D)', class Errors, trigger "O_Centror_AlarmW" bit 0
   1: 'Alarma stacker nou miscare verticala', class Errors, trigger "O_FurcaStacker_New_AlarmW" bit 3
   17: 'Furca stacker nu a coborat in timpul prestabilit (3D; S1_B3)', class Errors, trigger "O_Alm_Stack_Dwn" bit 0
   5: 'Alarma stacker miscare furci', class Errors, trigger "O_FurcaStacker_AlarmW" bit 3
   22: 'Furca stacker nou a pierdut detectia in pozitia retras (4D; S1_B13)', class Errors, trigger "O_FurcaStacker_New_AlarmW" bit 6
   11: 'Furca stacker nu s-a retras in timpul prestabilit (4D; S1_B13)', class Errors, trigger "O_FurcaStacker_AlarmW" bit 4
   3: 'Furca stacker nou blocata in pozitia de avans', class Errors, trigger "O_FurcaStacker_New_AlarmW" bit 5
   16: 'Furca stacker blocata in pozitia de jos', class Errors, trigger "O_Alm_Stack_Dwn" bit 1
   15: 'Furca stacker nu s-a ridicat in timpul prestabilit (3D; S1_B1)', class Errors, trigger "O_Alm_Stack_Up" bit 0
   6: 'Furcka stacker blocat in pozitia de avans', class Errors, trigger "O_FurcaStacker_AlarmW" bit 5
   14: 'Furca stacker a pierdut detectia in pozitia retras (4D; S1_B13)', class Errors, trigger "O_FurcaStacker_AlarmW" bit 6
   20: 'Furca stacker nou blocata in pozitia de retras', class Errors, trigger "O_FurcaStacker_New_AlarmW" bit 1
   57: 'Furca stacker a pierdut pozitia de sus (3D; S1_B1)', class Errors, trigger "O_Alm_Stack_Up" bit 2
   25: 'Centrorul a pierdut pozitia de retras (9D; CP2_SQ2)', class Errors, trigger "O_Centror_AlarmW" bit 6
   65: 'Furca stacker nou a pierdut pozitia de sus (3D; S1_B1)', class Errors, trigger "O_CilindruVerticalStacker_New_AlarmW" bit 2
   58: 'Furca stacker a pierdut pozitia de jos (3D; S1_B3)', class Errors, trigger "O_Alm_Stack_Dwn" bit 2
   63: 'Furca stacker nou nu s-a ridicat in timpul prestabilit (3D; S1_B1)', class Errors, trigger "O_CilindruVerticalStacker_New_AlarmW" bit 0
   62: 'Furca stacker nou nu a coborat in timpul prestabilit (3D; S1_B3)', class Errors, trigger "O_CilindruVerticalStacker_New_AlarmW" bit 4
   61: 'Furca stacker nou blocata in pozitia de jos', class Errors, trigger "O_CilindruVerticalStacker_New_AlarmW" bit 1
   64: 'Furca stacker nou a pierdut pozitia de jos (3D; S1_B3)', class Errors, trigger "O_CilindruVerticalStacker_New_AlarmW" bit 6
   23: 'Centrorul nu s-a retras in timpul prestabilit', class Errors, trigger "O_Centror_AlarmW" bit 4
   59: 'Furcka stacker blocata in pozitia de sus', class Errors, trigger "O_Alm_Stack_Up" bit 1
   60: 'Furcka stacker nou blocata in pozitia de sus', class Errors, trigger "O_CilindruVerticalStacker_New_AlarmW" bit 5
   24: 'Centrorul se afla in pozitia avans cu actionare', class Errors, trigger "O_Centror_AlarmW" bit 5
   66: 'General : Lipsa alimentare aer', class Errors, trigger "DB3_FAULTS_Alarm_General" bit 0
   67: 'Linia A : Lipsa aer stacker ch1', class Errors, trigger "DB3_FAULTS_Alarm_General" bit 1
   68: 'Linia B : Lipsa aer stacker nou ch1', class Errors, trigger "DB3_FAULTS_Alarm_General_SN" bit 1
   69: 'Linia A : Lipsa aer Z2_A ch1', class Errors, trigger "DB3_FAULTS_Alarm_General" bit 3
   72: 'Linia A : Lipsa power convertizor conveyor Staker -M3', class Errors, trigger "DB3_FAULTS_Alarm_General" bit 9
   73: 'Linia A : Lipsa power convertizor conveyor Staker -M4', class Errors, trigger "DB3_FAULTS_Alarm_General" bit 10
   74: 'Linia A : Lipsa aer Z2_A ch2', class Errors, trigger "DB3_FAULTS_Alarm_General" bit 6
   75: 'Linia B : Lipsa aer stacker nou ch2', class Errors, trigger "DB3_FAULTS_Alarm_General_SN" bit 4
   76: 'Linia A : Lipsa aer stacker ch2', class Errors, trigger "DB3_FAULTS_Alarm_General" bit 4
   77: 'Furca stacker nu a ajuns la mijloc in timpul prestabilit (3D; S1_B1)', class Errors, trigger "O_Alm_Stack_Mid" bit 0
   78: 'Furca stacker a pierdut pozitia de mijloc (3D; S1_B2)', class Errors, trigger "O_Alm_Stack_Mid" bit 2
   79: 'Furca stacker blocata in pozitia de mijloc(3D; S1_B2)', class Errors, trigger "O_Alm_Stack_Mid" bit 1
   47: 'Safety Linia B : Bariera mutting stacker dezarmata <111KF1>', class Errors, trigger "DB3_FAULTS_Alarm_Safety_SN" bit 3
   80: 'Linia B : Lipsa power convertizor conveyor Staker Nou -M2', class Errors, trigger "DB3_FAULTS_Alarm_General_SN" bit 10
   70: 'Linia B : Lipsa aer Z2_B ch1', class Errors, trigger "DB3_FAULTS_Alarm_General_SN" bit 3
   82: 'Linia B : Lipsa aer Z2_B ch2', class Errors, trigger "DB3_FAULTS_Alarm_General_SN" bit 6
   83: 'Linia B : Lipsa power convertizor conveyor Staker Nou -M1', class Errors, trigger "DB3_FAULTS_Alarm_General_SN" bit 9

text list "Text_list_1": 0 'Yes / Da'; 1 'No / Nu'; 2 ''; 3 ''; 4 ''

text list "Mod_Destacker": 1 'Energie'; 2 'Manual'; 3 'Asteptare Start'; 4 'Automat'; 5 'Init'; 5 'Safe'

text list "Mod_Stacker": 0 'Safe'; 1 'Energie'; 2 'Manual'; 3 'Asteptare Start'; 4 'Automat'; 5 'Init'

text list "Griper": 1 'retras'; 2 'avans'; 3 'spre av.'; 4 'spre ret.'; 5 'alarm'; 0 ''

text list "Palet": 0 'lipsa'; 1 'gol'; 2 'lucru'; 3 'plin'; 4 'alarm'

text list "sensCyl": 0 'avans'; 1 'retragere'; 2 'sus'; 3 'jos'

text list "msjOp_main": 1 'Alarma detectie produs pierduta la ppppppppppppp ,senzorul ssssssssss. Verificati daca produsul exista in fata senzorului e conform si bine asezat'

text list "numSenz": 0 'iCi'; 1 'iLa'; 2 'iLa_out'; 3 'iCm'; 4 'iCe'; 5 'iGrM'; 6 'iGrE'

